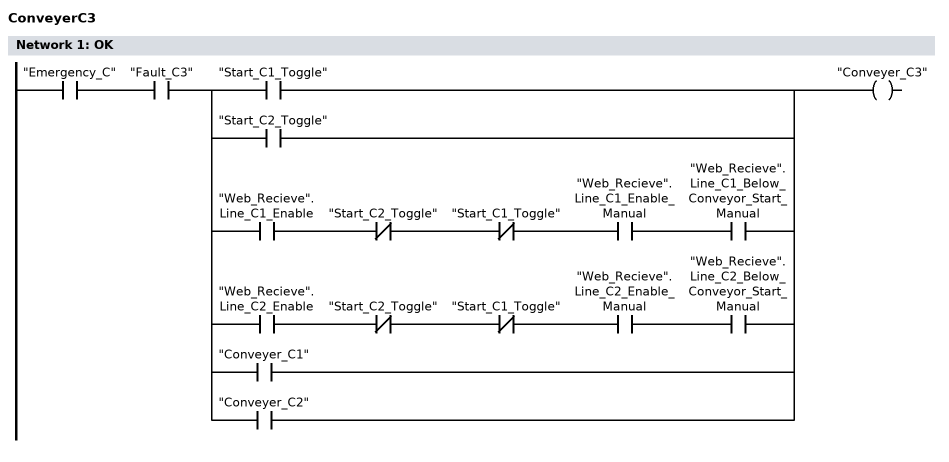
   RUNG wire#powerrail
      Contact( "Emergency_C" )
      Contact( "Fault_C3" )
      wire#w1
      Contact( "Start_C1_Toggle" )
      wire#w2
      Coil( "Conveyer_C3" )
   END_RUNG
   RUNG wire#w1
      Contact( "Start_C2_Toggle" )
   END_RUNG wire#w2
   RUNG wire#w1
      Contact( "Web_Recieve".Line_C1_Enable )
      I_Contact( "Start_C2_Toggle" )
      I_Contact( "Start_C1_Toggle" )
      Contact( "Web_Recieve".Line_C1_Enable_Manual )
      Contact( "Web_Recieve".Line_C1_Below_Conveyor_Start_Manual )
   END_RUNG wire#w2
   RUNG wire#w1
      Contact( "Web_Recieve".Line_C2_Enable )
      I_Contact( "Start_C2_Toggle" )
      I_Contact( "Start_C1_Toggle" )
      Contact( "Web_Recieve".Line_C2_Enable_Manual )
      Contact( "Web_Recieve".Line_C2_Below_Conveyor_Start_Manual )
   END_RUNG wire#w2
   RUNG wire#w1
      Contact( "Conveyer_C1" )
   END_RUNG wire#w2
   RUNG wire#w1
      Contact( "Conveyer_C2" )
   END_RUNG wire#w2
   // the same network as SCL:
   "Conveyer_C3" := "Emergency_C" AND "Fault_C3" AND ("Start_C1_Toggle" OR "Start_C2_Toggle" OR ("Web_Recieve".Line_C1_Enable AND NOT "Start_C2_Toggle" AND NOT "Start_C1_Toggle" AND "Web_Recieve".Line_C1_Enable_Manual AND "Web_Recieve".Line_C1_Below_Conveyor_Start_Manual) OR ("Web_Recieve".Line_C2_Enable AND NOT "Start_C2_Toggle" AND NOT "Start_C1_Toggle" AND "Web_Recieve".Line_C2_Enable_Manual AND "Web_Recieve".Line_C2_Below_Conveyor_Start_Manual) OR "Conveyer_C1" OR "Conveyer_C2");
END_REGION
END_FUNCTION_BLOCK

FUNCTION_BLOCK "WebDataPrepaare"   // FB10, SCL
{ S7_Optimized_Access := 'TRUE' }
VERSION : 0.1
BEGIN
   "Web_Send".C_Emergency := NOT "Emergency_C";
   "Web_Send".C1_Conveyer := "Conveyer_C1";
   "Web_Send".C2_Conveyer := "Conveyer_C2";
   "Web_Send".C3_Conveyor := "Conveyer_C3";

   "Web_Send".C1_Fault := NOT "Fault_C1";
   "Web_Send".C2_Fault := NOT "Fault_C2";
   "Web_Send".C3_Fault := NOT "Fault_C3";
   "Web_Send".C1_Silo_Low := "Low_Silo_C1";
   "Web_Send".C2_Silo_Low := "Low_Silo_C2";
   "Web_Send".C1_Silo_High := "HIgh_Silo_C1";
   "Web_Send".C2_Silo_High := "High_Silo_C2";
   "Web_Send".C1_Sample := "Pneumatic_C1";
   "Web_Send".C2_Sample := "Pneumatic_C2";
   "Web_Send".C1_Manual := "Web_Recieve".Line_C1_Enable_Manual;


   "Web_Send".C1_Running_Duration := "Web_Recieve".Line_C1_Conveyer_on_Time;
   "Web_Send".C1_Pause_Duration := "Web_Recieve".Line_C1_Conveyer_off_Time;
   "Web_Send".C1_Feeder_Vibration_Intensity := "Web_Recieve".Line_C1_Feeder_Intensity;
   "Web_Send".C1_Ruuning_Online := "Timer_On_C1_Conveyer".ET;
   "Web_Send".C1_Pause_Online := "Timer_Off_C1_Conveyer".ET;
   "Web_Send".C1_Sample_Interval :="Web_Recieve".Line_C1_Sampling_Time;
   "Web_Send".C1_Sample_Duration := "Web_Recieve".Line_C1_Sampling_OpenTime;
   "Web_Send".C1_Sample_Online := "Timer_Before_On_Sample_C1".ET - "Timer_Before_On_Sample_C1".ET;
   "Web_Send".C1_Enable := "Web_Recieve".Line_C1_Enable;
   "Web_Send".C1_Start := "Start_C1_Toggle";
   "Web_Send".C1_Empty_Line_Time := "Web_Recieve".Line_C1_Empty_Line_Time;
   "Web_Send".C1_Feeder_Delay_After_Start_Time := "Web_Recieve".Line_C1_Feeder_Delay_After_Start_Time;
   "Web_Send".C1_Feeder_Delay_Before_Stop_Time := "Web_Recieve".Line_C1_Feeder_Delay_Before_Stop_Time;
   "Web_Send".C1_Duration_Big_Silo_Stop_Time := "Web_Recieve".Line_C1_Big_Silo_Delay_Start;

   "Web_Send".C2_Running_Duration := "Web_Recieve".Line_C2_Conveyer_on_Time;
   "Web_Send".C2_Pause_Duration := "Web_Recieve".Line_C2_Conveyer_off_Time;
   "Web_Send".C2_Feeder_Vibration_Intensity := "Web_Recieve".Line_C2_Feeder_Intensity;
   "Web_Send".C2_Ruuning_Online := "Timer_On_C2_Conveyer".ET;
   "Web_Send".C2_Pause_Online := "Timer_Off_C2_Conveyer".ET;
   "Web_Send".C2_Sample_Interval := "Web_Recieve".Line_C2_Sampling_Time;
   "Web_Send".C2_Sample_Duration := "Web_Recieve".Line_C2_Sampling_OpenTime;
   "Web_Send".C2_Sample_Online := "Timer_Before_On_Sample_C2".ET - "Timer_Before_On_Sample_C2".ET;
   "Web_Send".C2_Enable := "Web_Recieve".Line_C2_Enable;
   "Web_Send".C2_Start := "Start_C2_Toggle";
   "Web_Send".C2_Empty_Line_Time := "Web_Recieve".Line_C2_Empty_Line_Time;
   "Web_Send".C2_Feeder_Delay_After_Start_Time := "Web_Recieve".Line_C2_Feeder_Delay_After_Start_Time;
   "Web_Send".C2_Feeder_Delay_Before_Stop_Time := "Web_Recieve".Line_C2_Feeder_Delay_Before_Stop_Time;
   "Web_Send".C2_Duration_Big_Silo_Stop_Time := "Web_Recieve".Line_C2_Big_Silo_Delay_Start;
END_FUNCTION_BLOCK

FUNCTION_BLOCK "Sample_C"   // FB11, LAD
{ S7_Optimized_Access := 'TRUE' }
VERSION : 0.1
   VAR_TEMP   // added for the SCL form of the ladder/FBD networks
      _w1 : Bool;
   END_VAR
BEGIN

REGION Network 1: C1 Before Sample
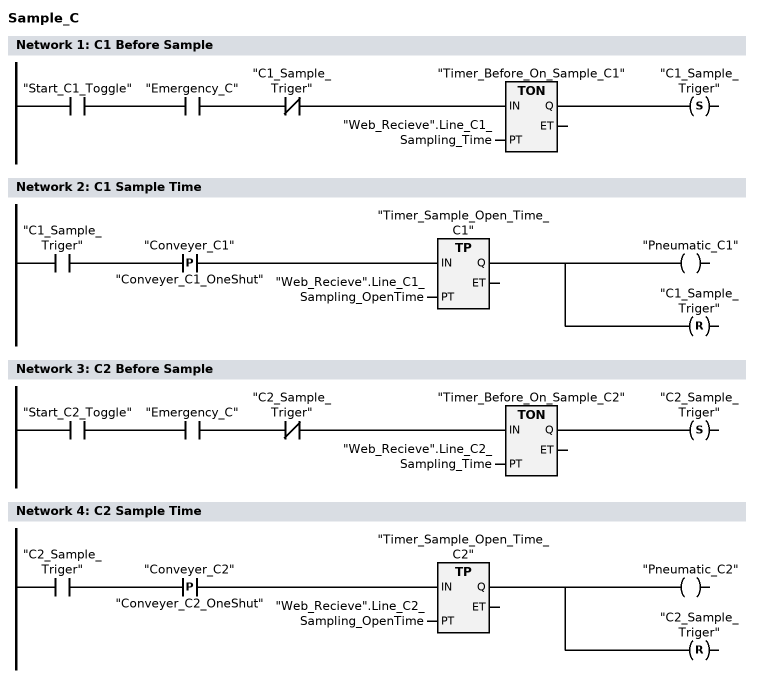
   "Timer_Before_On_Sample_C1".TON(IN := "Start_C1_Toggle" AND "Emergency_C" AND NOT "C1_Sample_Triger",
                           PT := "Web_Recieve".Line_C1_Sampling_Time);
   IF "Timer_Before_On_Sample_C1".Q THEN "C1_Sample_Triger" := TRUE; END_IF;
END_REGION

REGION Network 2: C1 Sample Time
   #_w1 := "C1_Sample_Triger" AND "Conveyer_C1" AND NOT "Conveyer_C1_OneShut";   // rising edge of "Conveyer_C1"
   "Conveyer_C1_OneShut" := "Conveyer_C1";
   "Timer_Sample_Open_Time_C1".TP(IN := #_w1, PT := "Web_Recieve".Line_C1_Sampling_OpenTime);
   "Pneumatic_C1" := "Timer_Sample_Open_Time_C1".Q;
   IF "Timer_Sample_Open_Time_C1".Q THEN "C1_Sample_Triger" := FALSE; END_IF;
END_REGION

REGION Network 3: C2 Before Sample
   "Timer_Before_On_Sample_C2".TON(IN := "Start_C2_Toggle" AND "Emergency_C" AND NOT "C2_Sample_Triger",
                           PT := "Web_Recieve".Line_C2_Sampling_Time);
   IF "Timer_Before_On_Sample_C2".Q THEN "C2_Sample_Triger" := TRUE; END_IF;
END_REGION

REGION Network 4: C2 Sample Time
   #_w1 := "C2_Sample_Triger" AND "Conveyer_C2" AND NOT "Conveyer_C2_OneShut";   // rising edge of "Conveyer_C2"
   "Conveyer_C2_OneShut" := "Conveyer_C2";
   "Timer_Sample_Open_Time_C2".TP(IN := #_w1, PT := "Web_Recieve".Line_C2_Sampling_OpenTime);
   "Pneumatic_C2" := "Timer_Sample_Open_Time_C2".Q;
   IF "Timer_Sample_Open_Time_C2".Q THEN "C2_Sample_Triger" := FALSE; END_IF;
END_REGION
END_FUNCTION_BLOCK

FUNCTION_BLOCK "Silo_Big_C"   // FB12, LAD
{ S7_Optimized_Access := 'TRUE' }
VERSION : 0.1
BEGIN

REGION Network 1
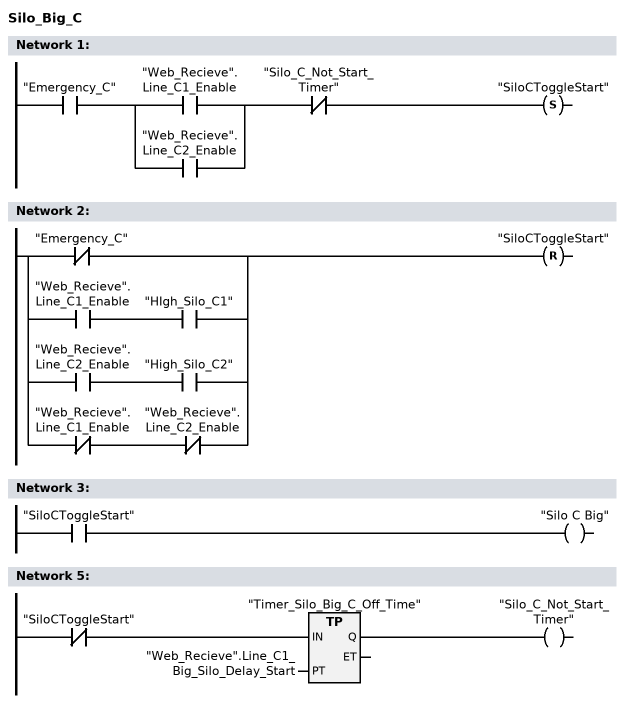
   RUNG wire#powerrail
      Contact( "Emergency_C" )
      wire#w1
      Contact( "Web_Recieve".Line_C1_Enable )
      wire#w2
      I_Contact( "Silo_C_Not_Start_Timer" )
      S_Coil( "SiloCToggleStart" )
   END_RUNG
   RUNG wire#w1
      Contact( "Web_Recieve".Line_C2_Enable )
   END_RUNG wire#w2
   // the same network as SCL:
   IF "Emergency_C" AND ("Web_Recieve".Line_C1_Enable OR "Web_Recieve".Line_C2_Enable) AND NOT "Silo_C_Not_Start_Timer" THEN
       "SiloCToggleStart" := TRUE;
   END_IF;
END_REGION

REGION Network 2
   RUNG wire#powerrail
      I_Contact( "Emergency_C" )
      wire#w1
      R_Coil( "SiloCToggleStart" )
   END_RUNG
   RUNG wire#powerrail
      Contact( "Web_Recieve".Line_C1_Enable )
      Contact( "HIgh_Silo_C1" )
   END_RUNG wire#w1
   RUNG wire#powerrail
      Contact( "Web_Recieve".Line_C2_Enable )
      Contact( "High_Silo_C2" )
   END_RUNG wire#w1
   RUNG wire#powerrail
      I_Contact( "Web_Recieve".Line_C1_Enable )
      I_Contact( "Web_Recieve".Line_C2_Enable )
   END_RUNG wire#w1
   // the same network as SCL:
   IF NOT "Emergency_C" OR ("Web_Recieve".Line_C1_Enable AND "HIgh_Silo_C1") OR ("Web_Recieve".Line_C2_Enable AND "High_Silo_C2") OR (NOT "Web_Recieve".Line_C1_Enable AND NOT "Web_Recieve".Line_C2_Enable) THEN
       "SiloCToggleStart" := FALSE;
   END_IF;
END_REGION

REGION Network 3
   RUNG wire#powerrail
      Contact( "SiloCToggleStart" )
      Coil( "Silo C Big" )
   END_RUNG
   // the same network as SCL:
   "Silo C Big" := "SiloCToggleStart";
END_REGION

REGION Network 5
   "Timer_Silo_Big_C_Off_Time".TP(IN := NOT "SiloCToggleStart",
                           PT := "Web_Recieve".Line_C1_Big_Silo_Delay_Start);
   "Silo_C_Not_Start_Timer" := "Timer_Silo_Big_C_Off_Time".Q;
END_REGION
END_FUNCTION_BLOCK

FUNCTION_BLOCK "Empty Line C1"   // FB13, LAD
{ S7_Optimized_Access := 'TRUE' }
VERSION : 0.1
BEGIN

REGION Network 1
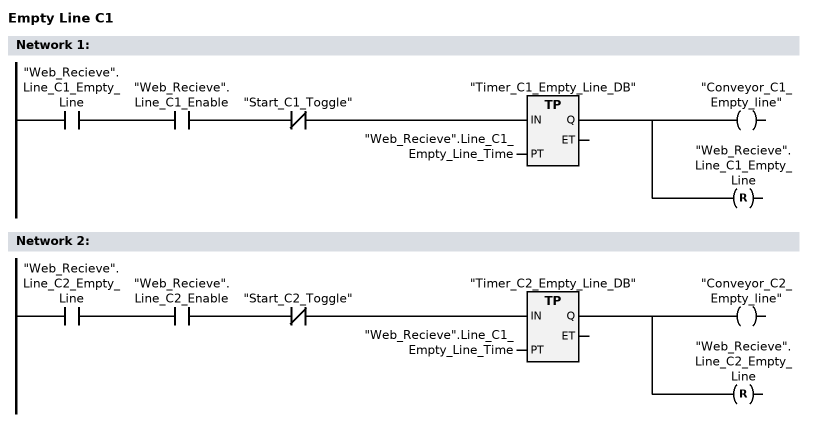
   "Timer_C1_Empty_Line_DB".TP(IN := "Web_Recieve".Line_C1_Empty_Line AND "Web_Recieve".Line_C1_Enable AND NOT "Start_C1_Toggle",
                           PT := "Web_Recieve".Line_C1_Empty_Line_Time);
   "Conveyor_C1_Empty_line" := "Timer_C1_Empty_Line_DB".Q;
   IF "Timer_C1_Empty_Line_DB".Q THEN "Web_Recieve".Line_C1_Empty_Line := FALSE; END_IF;
END_REGION

REGION Network 2
   "Timer_C2_Empty_Line_DB".TP(IN := "Web_Recieve".Line_C2_Empty_Line AND "Web_Recieve".Line_C2_Enable AND NOT "Start_C2_Toggle",
                           PT := "Web_Recieve".Line_C1_Empty_Line_Time);
   "Conveyor_C2_Empty_line" := "Timer_C2_Empty_Line_DB".Q;
   IF "Timer_C2_Empty_Line_DB".Q THEN "Web_Recieve".Line_C2_Empty_Line := FALSE; END_IF;
END_REGION
END_FUNCTION_BLOCK

ORGANIZATION_BLOCK "Main"   // OB1, LAD, ProgramCycle
TITLE = "Main Program Sweep (Cycle)"
{ S7_Optimized_Access := 'TRUE' }
VERSION : 0.1
   VAR_INPUT
      Initial_Call : Bool;   // Initial call of this OB
      Remanence : Bool;   // =True, if remanent data are available
   END_VAR
   VAR_TEMP
      TEMP : Int;
      clkRetVal : Int;
      newt : Int;
   END_VAR
BEGIN

REGION Network 1
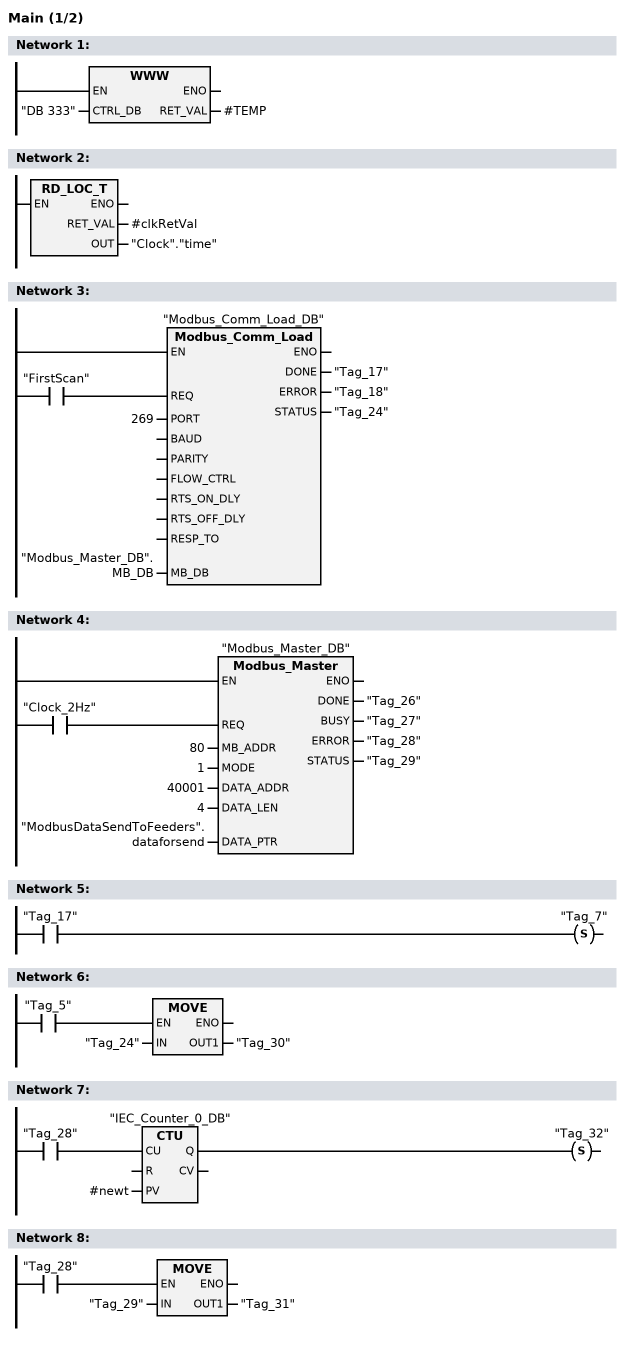
   #TEMP := WWW(CTRL_DB := "DB 333");
END_REGION

REGION Network 2
   #clkRetVal := RD_LOC_T(OUT => "Clock"."time");
END_REGION

REGION Network 3
   "Modbus_Comm_Load_DB"(REQ := "FirstScan",   // Modbus_Comm_Load
                         PORT := 269,
                         MB_DB := "Modbus_Master_DB".MB_DB,
                         DONE => "Tag_17",
                         ERROR => "Tag_18",
                         STATUS => "Tag_24");
END_REGION

REGION Network 4
   "Modbus_Master_DB"(REQ := "Clock_2Hz",   // Modbus_Master
                      MB_ADDR := 80,
                      MODE := 1,
                      DATA_ADDR := 40001,
                      DATA_LEN := 4,
                      DATA_PTR := "ModbusDataSendToFeeders".dataforsend,
                      DONE => "Tag_26",
                      BUSY => "Tag_27",
                      ERROR => "Tag_28",
                      STATUS => "Tag_29");
END_REGION

REGION Network 5
   RUNG wire#powerrail
      Contact( "Tag_17" )
      S_Coil( "Tag_7" )
   END_RUNG
   // the same network as SCL:
   IF "Tag_17" THEN "Tag_7" := TRUE; END_IF;
END_REGION

REGION Network 6
   RUNG wire#powerrail
      Contact( "Tag_5" )
      Move(in := "Tag_24", out1 => "Tag_30")
   END_RUNG
   // the same network as SCL:
   IF "Tag_5" THEN "Tag_30" := "Tag_24"; END_IF;
END_REGION

REGION Network 7
   "IEC_Counter_0_DB".CTU(CU := "Tag_28", PV := #newt);
   IF "IEC_Counter_0_DB".Q THEN "Tag_32" := TRUE; END_IF;
END_REGION

REGION Network 8
   RUNG wire#powerrail
      Contact( "Tag_28" )
      Move(in := "Tag_29", out1 => "Tag_31")
   END_RUNG
   // the same network as SCL:
   IF "Tag_28" THEN "Tag_31" := "Tag_29"; END_IF;
END_REGION

REGION Network 9
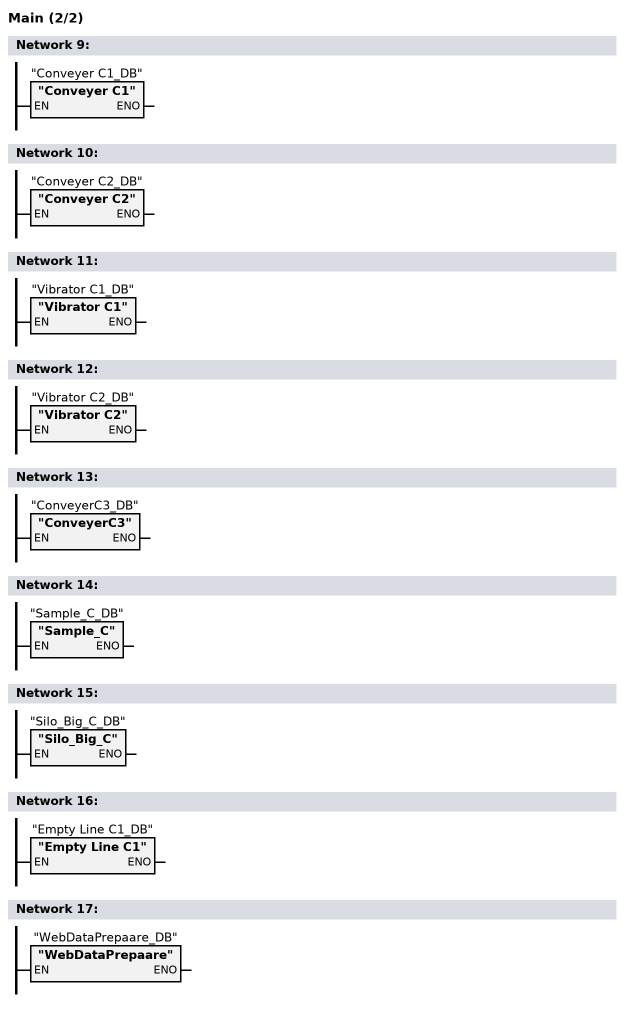
   RUNG wire#powerrail
      "Conveyer C1_DB"()
   END_RUNG
   // the same network as SCL:
   "Conveyer C1_DB"();   // "Conveyer C1"
END_REGION

REGION Network 10
   RUNG wire#powerrail
      "Conveyer C2_DB"()
   END_RUNG
   // the same network as SCL:
   "Conveyer C2_DB"();   // "Conveyer C2"
END_REGION

REGION Network 11
   RUNG wire#powerrail
      "Vibrator C1_DB"()
   END_RUNG
   // the same network as SCL:
   "Vibrator C1_DB"();   // "Vibrator C1"
END_REGION

REGION Network 12
   RUNG wire#powerrail
      "Vibrator C2_DB"()
   END_RUNG
   // the same network as SCL:
   "Vibrator C2_DB"();   // "Vibrator C2"
END_REGION

REGION Network 13
   RUNG wire#powerrail
      "ConveyerC3_DB"()
   END_RUNG
   // the same network as SCL:
   "ConveyerC3_DB"();   // "ConveyerC3"
END_REGION

REGION Network 14
   RUNG wire#powerrail
      "Sample_C_DB"()
   END_RUNG
   // the same network as SCL:
   "Sample_C_DB"();   // "Sample_C"
END_REGION

REGION Network 15
   RUNG wire#powerrail
      "Silo_Big_C_DB"()
   END_RUNG
   // the same network as SCL:
   "Silo_Big_C_DB"();   // "Silo_Big_C"
END_REGION

REGION Network 16
   RUNG wire#powerrail
      "Empty Line C1_DB"()
   END_RUNG
   // the same network as SCL:
   "Empty Line C1_DB"();   // "Empty Line C1"
END_REGION

REGION Network 17
   RUNG wire#powerrail
      "WebDataPrepaare_DB"()
   END_RUNG
   // the same network as SCL:
   "WebDataPrepaare_DB"();   // "WebDataPrepaare"
END_REGION
END_ORGANIZATION_BLOCK

// ===== PLC "PLC_1"  CPU 1516-3 PN/DP =====

VAR_GLOBAL   // PLC tag table "Default tag table"
   "Tag_31" AT %M100.5 : Bool;
   "Run consent OS" AT %M151.6 : Bool;
   "Run_Consent_A1_Negetive_OS" AT %M151.7 : Bool;
   "Vibrator_A2_Remaning_Time" AT %MD166 : DInt;
   "System_Byte(1)" AT %MB1 : Byte;
   "FirstScan" AT %M1.0 : Bool;
END_VAR

VAR_GLOBAL   // PLC tag table "Default tag table_1"
   "Phase_Control" AT %I8.0 : Bool;
   "Start_A" AT %I8.7 : Bool;
   "Spare_6" AT %I9.6 : Bool;
   "Spare_7" AT %I9.7 : Bool;
   "Emergency_A" AT %I8.4 : Bool;
   "Fault_A1" AT %I8.1 : Bool;
   "Low_Silo_A1" AT %I0.2 : Bool;
   "Low_Silo_A2" AT %I0.1 : Bool;
   "Low_Silo_B1" AT %I0.7 : Bool;
   "Low_Silo_B2" AT %I0.4 : Bool;
   "High_Silo_A1" AT %I0.3 : Bool;
   "High_Silo_A2" AT %I0.0 : Bool;
   "High_Silo_B1" AT %I0.6 : Bool;
   "High_Silo_B2" AT %I0.5 : Bool;
   "Fault_A2" AT %I9.1 : Bool;
   "Fault_B1" AT %I8.2 : Bool;
   "Fault_B2" AT %I9.2 : Bool;
   "Fault_A3" AT %I9.5 : Bool;
   "Fault_B3" AT %I9.4 : Bool;
   "Emergency_B" AT %I9.3 : Bool;
   "Rel Spare_4" AT %Q2.4 : Bool;
   "Rel Spare_5" AT %Q2.5 : Bool;
   "Rel Spare_6" AT %Q2.6 : Bool;
   "Rel Spare_7" AT %Q2.7 : Bool;
   "Rel Spare_8" AT %Q3.0 : Bool;
   "Rel Spare_9" AT %Q3.1 : Bool;
   "Rel Spare_10" AT %Q3.2 : Bool;
   "Rel Spare_11" AT %Q3.3 : Bool;
   "Rel Spare_12" AT %Q3.4 : Bool;
   "Rel Spare_13" AT %Q3.5 : Bool;
   "Rel Spare_14" AT %Q3.6 : Bool;
   "Rel Spare_15" AT %Q3.7 : Bool;
   "Light_A1" AT %Q2.3 : Bool;
   "Light_A2" AT %Q2.2 : Bool;
   "Light_B1" AT %Q2.1 : Bool;
   "Light_B2" AT %Q2.0 : Bool;
   "Conveyer_A1" AT %Q0.4 : Bool;
   "Conveyer_A2" AT %Q0.5 : Bool;
   "Conveyer_B1" AT %Q9.0 : Bool;
   "Conveyer_B2" AT %Q8.0 : Bool;
   "Pneumatic_A1" AT %Q9.1 : Bool;
   "Pneumatic_A2" AT %Q8.1 : Bool;
   "Pneumatic_B1" AT %Q8.2 : Bool;
   "Pneumatic_B2" AT %Q9.2 : Bool;
   "Conveyer_A3" AT %Q9.5 : Bool;
   "Conveyer_B3_Left" AT %Q9.6 : Bool;
   "Conveyer_B3_Right" AT %Q8.5 : Bool;
   "Tag_1(1)" AT %M10.0 : Bool;
   "Tag_2" AT %M10.1 : Bool;
   "start" AT %M10.2 : Bool;
   "Tag_3" AT %M110.0 : Bool;
   "Tag_10" AT %M110.1 : Bool;
   "Tag_11" AT %M110.2 : Bool;
   "System_Byte" AT %MB1 : Byte;
   "DiagStatusUpdate" AT %M1.1 : Bool;
   "AlwaysTRUE" AT %M1.2 : Bool;
   "AlwaysFALSE" AT %M1.3 : Bool;
   "Clock_Byte" AT %MB0 : Byte;
   "Clock_10Hz" AT %M0.0 : Bool;
   "Clock_5Hz" AT %M0.1 : Bool;
   "Clock_2.5Hz" AT %M0.2 : Bool;
   "Clock_2Hz" AT %M0.3 : Bool;
   "Clock_1.25Hz" AT %M0.4 : Bool;
   "Clock_1Hz" AT %M0.5 : Bool;
   "Clock_0.625Hz" AT %M0.6 : Bool;
   "Clock_0.5Hz" AT %M0.7 : Bool;
   "Tag_12" AT %M120.1 : Bool;
   "Tag_13" AT %M120.0 : Bool;
   "Tag_14" AT %M120.2 : Bool;
   "Tag_15" AT %MW112 : Word;
   "Tag_16" AT %MW114 : Word;
   "Tag_17" AT %MW122 : Word;
   "Tag_18" AT %MW124 : Word;
   "Tag_4" AT %M1000.0 : Bool;
   "Tag_5" AT %M1000.1 : Bool;
   "Tag_6" AT %MW1002 : Word;
   "Tag_7" AT %M1000.4 : Bool;
   "Tag_8" AT %MW1004 : Word;
   "Tag_9" AT %M1010.0 : Bool;
   "Tag_19" AT %M1010.1 : Bool;
   "Tag_20" AT %M1010.2 : Bool;
   "Tag_21" AT %MW1012 : Word;
   "Tag_22" AT %M1010.4 : Bool;
   "Tag_23" AT %MW1014 : Word;
   "Tag_24" AT %M990.0 : Bool;
   "Tag_25" AT %M990.5 : Bool;
   "Line_A1_Start_Consent" AT %M150.0 : Bool;
   "Line_A1_Run_Consent" AT %M150.1 : Bool;
   "Line_A1_Conveyer_Timer" AT %M150.2 : Bool;
   "A1_Start_Conveyer" AT %M150.3 : Bool;
   "TriggerStartToggleMemory" AT %M150.4 : Bool;
   "Start_A1_Toggle" AT %M150.5 : Bool;
   "TriggerA1ToggleStop" AT %M150.6 : Bool;
   "Conveyer_A1_On" AT %M150.7 : Bool;
   "Conveyer_A1_Off" AT %M151.0 : Bool;
   "Line_A2_Start_Consent" AT %M160.0 : Bool;
   "Line_A2_Run_Consent" AT %M160.1 : Bool;
   "Line_A2_Conveyer_Timer" AT %M160.2 : Bool;
   "A2_Start_Conveyer" AT %M160.3 : Bool;
   "TriggerStopToggleMemoryA2" AT %M160.6 : Bool;
   "TriggerStartToggleMemoryA2" AT %M160.4 : Bool;
   "Start_A2_Toggle" AT %M160.5 : Bool;
   "Conveyer_A2_Off" AT %M161.0 : Bool;
   "Conveyer_A2_On" AT %M160.7 : Bool;
   "Line_B1_Start_Consent" AT %M170.0 : Bool;
   "Line_B1_Run_Consent" AT %M170.1 : Bool;
   "Line_B1_Conveyer_Timer" AT %M170.2 : Bool;
   "B1_Start_Conveyer" AT %M170.3 : Bool;
   "Start_B1_Toggle" AT %M170.5 : Bool;
   "TriggerStartToggleMemoryB1" AT %M170.4 : Bool;
   "TriggerB1ToggleStop" AT %M170.6 : Bool;
   "Conveyer_B1_Off" AT %M171.0 : Bool;
   "Conveyer_B1_On" AT %M170.7 : Bool;
   "Line_B2_Start_Consent" AT %M180.0 : Bool;
   "Line_B2_Run_Consent" AT %M180.1 : Bool;
   "B2_Start_Conveyer" AT %M180.3 : Bool;
   "Line_B2_Conveyer_Timer" AT %M180.2 : Bool;
   "Start_B2_Toggle" AT %M180.5 : Bool;
   "TriggerStartToggleMemoryB2" AT %M180.4 : Bool;
   "TriggerStopToggleMemoryB2" AT %M180.6 : Bool;
   "Conveyer_B2_Off" AT %M181.0 : Bool;
   "Conveyer_B2_On" AT %M180.7 : Bool;
   "Vibrator_A1_On" AT %M151.4 : Bool;
   "Vibrator_A2_On" AT %M161.4 : Bool;
   "Vibrator_B1_On" AT %M171.4 : Bool;
   "Vibrator_B2_On" AT %M181.4 : Bool;
   "A1_Sample_Triger" AT %M151.1 : Bool;
   "Conveyer_A1_OneShut" AT %M151.2 : Bool;
   "Tag_27" AT %M151.3 : Bool;
   "A2_Sample_Triger" AT %M161.1 : Bool;
   "Conveyer_A2_OneShut" AT %M161.2 : Bool;
   "B1_Sample_Triger" AT %M171.1 : Bool;
   "Conveyer_B1_OneShut" AT %M171.2 : Bool;
   "B2_Sample_Triger" AT %M181.1 : Bool;
   "Conveyer_B2_OneShut" AT %M181.2 : Bool;
   "B_Emergency_Flag" AT %M171.3 : Bool;
   "SiloAToggleStart" AT %M190.0 : Bool;
   "SiloBToggleStart" AT %M190.1 : Bool;
   "Conveyor_B3_Left" AT %M200.0 : Bool;
   "Conveyor_B3_Right" AT %M200.1 : Bool;
   "Silo_B_Not_Start_Timer" AT %M190.3 : Bool;
   "Silo_A_Not_Start_Timer" AT %M190.2 : Bool;
   "Conveyor_B3_Start" AT %M190.4 : Bool;
   "Conveyor_A1_Empty_line" AT %M151.5 : Bool;
   "Conveyor_A2_Empty_line" AT %M161.5 : Bool;
   "Conveyor_B1_Empty_line" AT %M171.5 : Bool;
   "Conveyor_B2_Empty_line" AT %M181.5 : Bool;
   "Vibrator_A1_Remaning_Time" AT %MD156 : DInt;
   "Tag_29" AT %MD176 : DInt;
   "Tag_30" AT %MD186 : DInt;
END_VAR

VAR_GLOBAL CONSTANT   // PLC tag table "Default tag table_1"
   "None(1)" : Pip := 65535;
   "Automatic update(1)" : Pip := 0;
   "PIP 1(1)" : Pip := 1;
   "PIP 2(1)" : Pip := 2;
   "PIP 3(1)" : Pip := 3;
   "PIP 4(1)" : Pip := 4;
   "PIP OB Servo(1)" : Pip := 32768;
   "Local~MC(1)" : Hw_SubModule := 51;
   "Local~Common(1)" : Hw_SubModule := 50;
   "Local~Device(1)" : Hw_Device := 32;
   "Local~Configuration(1)" : Hw_SubModule := 33;
   "Local~Exec(1)" : Hw_SubModule := 52;
   "Local(1)" : Hw_SubModule := 49;
   "Local~PROFINET_interface_1(1)" : Hw_Interface := 64;
   "Local~PROFINET_interface_1~Port_1(1)" : Hw_Interface := 65;
   "Local~HSC_1" : Hw_Hsc := 257;
   "Local~HSC_2" : Hw_Hsc := 258;
   "Local~HSC_3" : Hw_Hsc := 259;
   "Local~HSC_4" : Hw_Hsc := 260;
   "Local~HSC_5" : Hw_Hsc := 261;
   "Local~HSC_6" : Hw_Hsc := 262;
   "Local~AI_2_1" : Hw_SubModule := 263;
   "Local~DI_8_DQ_6_1" : Hw_SubModule := 264;
   "Local~Pulse_1" : Hw_Pwm := 265;
   "Local~Pulse_2" : Hw_Pwm := 266;
   "Local~Pulse_3" : Hw_Pwm := 267;
   "Local~Pulse_4" : Hw_Pwm := 268;
   "Local~CB_1241_(RS485)" : Port := 269;
   "Local~DQ_16xRelay_1" : Hw_SubModule := 270;
   "Local~DI_16x24VDC_DQ_16xRelay_1" : Hw_SubModule := 271;
   "OB_Main(1)" : OB_PCYCLE := 1;
END_VAR

DATA_BLOCK "ScenarioData"   // DB1
{ S7_Optimized_Access := 'TRUE' }
VERSION : 0.1
   VAR
      DefaultScenario : Int := 1;
      Line_A1_Conveyer_on_Time_Scenario_A : DInt := 2;
      Line_A1_Conveyer_off_Time_Scenario_A : DInt := 3;
      Line_A1_Sampling_Time_Scenario_A : DInt := 4;
      Line_A1_Sampling_OpenTime_Scenario_A : DInt := 5;
      Line_A1_Feeder_Intensity_Scenario_A : Int := 6;
      Line_A1_Duration_Big_Silo_Off_Scenario_A : DInt := 7;
      Line_A1_Feeder_Delay_Before_Stop_Time_Scenario_A : DInt := 8;
      Line_A1_Feeder_Delay_After_Start_Time_Scenario_A : DInt := 9;
      Line_A1_Conveyer_on_Time_Scenario_B : DInt := 10;
      Line_A1_Conveyer_off_Time_Scenario_B : DInt := 11;
      Line_A1_Sampling_Time_Scenario_B : DInt := 12;
      Line_A1_Sampling_OpenTime_Scenario_B : DInt := 13;
      Line_A1_Feeder_Intensity_Scenario_B : Int := 14;
      Line_A1_Duration_Big_Silo_Off_Scenario_B : DInt := 15;
      Line_A1_Feeder_Delay_Before_Stop_Time_Scenario_B : DInt := 16;
      Line_A1_Feeder_Delay_After_Start_Time_Scenario_B : DInt := 17;
      Line_A1_Conveyer_on_Time_Scenario_C : DInt := 18;
      Line_A1_Conveyer_off_Time_Scenario_C : DInt := 19;
      Line_A1_Sampling_Time_Scenario_C : DInt := 20;
      Line_A1_Sampling_OpenTime_Scenario_C : DInt := 21;
      Line_A1_Feeder_Intensity_Scenario_C : Int := 22;
      Line_A1_Duration_Big_Silo_Off_Scenario_C : DInt := 23;
      Line_A1_Feeder_Delay_Before_Stop_Time_Scenario_C : DInt := 24;
      Line_A1_Feeder_Delay_After_Start_Time_Scenario_C : DInt := 25;
      Line_A1_Conveyer_on_Time_Scenario_E : DInt := 26;
      Line_A1_Conveyer_off_Time_Scenario_E : DInt := 27;
      Line_A1_Sampling_Time_Scenario_E : DInt := 28;
      Line_A1_Sampling_OpenTime_Scenario_E : DInt := 29;
      Line_A1_Feeder_Intensity_Scenario_E : Int := 30;
      Line_A1_Duration_Big_Silo_Off_Scenario_E : DInt := 31;
      Line_A1_Feeder_Delay_Before_Stop_Time_Scenario_E : DInt := 32;
      Line_A1_Feeder_Delay_After_Start_Time_Scenario_E : DInt := 33;
      Line_A1_Conveyer_on_Time_Scenario_D : DInt := 34;
      Line_A1_Conveyer_off_Time_Scenario_D : DInt := 35;
      Line_A1_Sampling_Time_Scenario_D : DInt := 36;
      Line_A1_Sampling_OpenTime_Scenario_D : DInt := 37;
      Line_A1_Feeder_Intensity_Scenario_D : Int := 38;
      Line_A1_Duration_Big_Silo_Off_Scenario_D : DInt := 39;
      Line_A1_Feeder_Delay_Before_Stop_Time_Scenario_D : DInt := 40;
      Line_A1_Feeder_Delay_After_Start_Time_Scenario_D : DInt := 41;
      Line_A2_Conveyer_on_Time_Scenario_A : DInt := 42;
      Line_A2_Conveyer_off_Time_Scenario_A : DInt := 43;
      Line_A2_Sampling_Time_Scenario_A : DInt := 44;
      Line_A2_Sampling_OpenTime_Scenario_A : DInt := 45;
      Line_A2_Feeder_Intensity_Scenario_A : Int := 46;
      Line_A2_Duration_Big_Silo_Off_Scenario_A : DInt := 47;
      Line_A2_Feeder_Delay_Before_Stop_Time_Scenario_A : DInt := 48;
      Line_A2_Feeder_Delay_After_Start_Time_Scenario_A : DInt := 49;
      Line_A2_Conveyer_on_Time_Scenario_B : DInt := 50;
      Line_A2_Conveyer_off_Time_Scenario_B : DInt := 51;
      Line_A2_Sampling_Time_Scenario_B : DInt := 52;
      Line_A2_Sampling_OpenTime_Scenario_B : DInt := 53;
      Line_A2_Feeder_Intensity_Scenario_B : Int := 54;
      Line_A2_Duration_Big_Silo_Off_Scenario_B : DInt := 55;
      Line_A2_Feeder_Delay_Before_Stop_Time_Scenario_B : DInt := 56;
      Line_A2_Feeder_Delay_After_Start_Time_Scenario_B : DInt := 57;
      Line_A2_Conveyer_on_Time_Scenario_C : DInt := 58;
      Line_A2_Conveyer_off_Time_Scenario_C : DInt := 59;
      Line_A2_Sampling_Time_Scenario_C : DInt := 60;
      Line_A2_Sampling_OpenTime_Scenario_C : DInt := 61;
      Line_A2_Feeder_Intensity_Scenario_C : Int := 62;
      Line_A2_Duration_Big_Silo_Off_Scenario_C : DInt := 63;
      Line_A2_Feeder_Delay_Before_Stop_Time_Scenario_C : DInt := 64;
      Line_A2_Feeder_Delay_After_Start_Time_Scenario_C : DInt := 65;
      Line_A2_Conveyer_on_Time_Scenario_E : DInt := 66;
      Line_A2_Conveyer_off_Time_Scenario_E : DInt := 67;
      Line_A2_Sampling_Time_Scenario_E : DInt := 68;
      Line_A2_Sampling_OpenTime_Scenario_E : DInt := 69;
      Line_A2_Feeder_Intensity_Scenario_E : Int := 70;
      Line_A2_Duration_Big_Silo_Off_Scenario_E : DInt := 71;
      Line_A2_Feeder_Delay_Before_Stop_Time_Scenario_E : DInt := 72;
      Line_A2_Feeder_Delay_After_Start_Time_Scenario_E : DInt := 73;
      Line_A2_Conveyer_on_Time_Scenario_D : DInt := 74;
      Line_A2_Conveyer_off_Time_Scenario_D : DInt := 75;
      Line_A2_Sampling_Time_Scenario_D : DInt := 76;
      Line_A2_Sampling_OpenTime_Scenario_D : DInt := 77;
      Line_A2_Feeder_Intensity_Scenario_D : Int := 78;
      Line_A2_Duration_Big_Silo_Off_Scenario_D : DInt := 79;
      Line_A2_Feeder_Delay_Before_Stop_Time_Scenario_D : DInt := 80;
      Line_A2_Feeder_Delay_After_Start_Time_Scenario_D : DInt := 81;
      Line_B1_Conveyer_on_Time_Scenario_A : DInt := 82;
      Line_B1_Conveyer_off_Time_Scenario_A : DInt := 83;
      Line_B1_Sampling_Time_Scenario_A : DInt := 84;
      Line_B1_Sampling_OpenTime_Scenario_A : DInt := 85;
      Line_B1_Feeder_Intensity_Scenario_A : Int := 86;
      Line_B1_Duration_Big_Silo_Off_Scenario_A : DInt := 87;
      Line_B1_Feeder_Delay_Before_Stop_Time_Scenario_A : DInt := 88;
      Line_B1_Feeder_Delay_After_Start_Time_Scenario_A : DInt := 89;
      Line_B1_Conveyer_on_Time_Scenario_B : DInt := 90;
      Line_B1_Conveyer_off_Time_Scenario_B : DInt := 91;
      Line_B1_Sampling_Time_Scenario_B : DInt := 92;
      Line_B1_Sampling_OpenTime_Scenario_B : DInt := 93;
      Line_B1_Feeder_Intensity_Scenario_B : Int := 94;
      Line_B1_Duration_Big_Silo_Off_Scenario_B : DInt := 95;
      Line_B1_Feeder_Delay_Before_Stop_Time_Scenario_B : DInt := 96;
      Line_B1_Feeder_Delay_After_Start_Time_Scenario_B : DInt := 97;
      Line_B1_Conveyer_on_Time_Scenario_C : DInt := 98;
      Line_B1_Conveyer_off_Time_Scenario_C : DInt := 99;
      Line_B1_Sampling_Time_Scenario_C : DInt := 100;
      Line_B1_Sampling_OpenTime_Scenario_C : DInt := 101;
      Line_B1_Feeder_Intensity_Scenario_C : Int := 102;
      Line_B1_Duration_Big_Silo_Off_Scenario_C : DInt := 103;
      Line_B1_Feeder_Delay_Before_Stop_Time_Scenario_C : DInt := 104;
      Line_B1_Feeder_Delay_After_Start_Time_Scenario_C : DInt := 105;
      Line_B1_Conveyer_on_Time_Scenario_E : DInt := 106;
      Line_B1_Conveyer_off_Time_Scenario_E : DInt := 107;
      Line_B1_Sampling_Time_Scenario_E : DInt := 108;
      Line_B1_Sampling_OpenTime_Scenario_E : DInt := 109;
      Line_B1_Feeder_Intensity_Scenario_E : Int := 110;
      Line_B1_Duration_Big_Silo_Off_Scenario_E : DInt := 111;
      Line_B1_Feeder_Delay_Before_Stop_Time_Scenario_E : DInt := 112;
      Line_B1_Feeder_Delay_After_Start_Time_Scenario_E : DInt := 113;
      Line_B1_Conveyer_on_Time_Scenario_D : DInt := 114;
      Line_B1_Conveyer_off_Time_Scenario_D : DInt := 115;
      Line_B1_Sampling_Time_Scenario_D : DInt := 116;
      Line_B1_Sampling_OpenTime_Scenario_D : DInt := 117;
      Line_B1_Feeder_Intensity_Scenario_D : Int := 118;
      Line_B1_Duration_Big_Silo_Off_Scenario_D : DInt := 119;
      Line_B1_Feeder_Delay_Before_Stop_Time_Scenario_D : DInt := 120;
      Line_B1_Feeder_Delay_After_Start_Time_Scenario_D : DInt := 121;
      Line_B2_Conveyer_on_Time_Scenario_A : DInt := 122;
      Line_B2_Conveyer_off_Time_Scenario_A : DInt := 123;
      Line_B2_Sampling_Time_Scenario_A : DInt := 124;
      Line_B2_Sampling_OpenTime_Scenario_A : DInt := 125;
      Line_B2_Feeder_Intensity_Scenario_A : Int := 126;
      Line_B2_Duration_Big_Silo_Off_Scenario_A : DInt := 127;
      Line_B2_Feeder_Delay_Before_Stop_Time_Scenario_A : DInt := 128;
      Line_B2_Feeder_Delay_After_Start_Time_Scenario_A : DInt := 129;
      Line_B2_Conveyer_on_Time_Scenario_B : DInt := 130;
      Line_B2_Conveyer_off_Time_Scenario_B : DInt := 131;
      Line_B2_Sampling_Time_Scenario_B : DInt := 132;
      Line_B2_Sampling_OpenTime_Scenario_B : DInt := 133;
      Line_B2_Feeder_Intensity_Scenario_B : Int := 134;
      Line_B2_Duration_Big_Silo_Off_Scenario_B : DInt := 135;
      Line_B2_Feeder_Delay_Before_Stop_Time_Scenario_B : DInt := 136;
      Line_B2_Feeder_Delay_After_Start_Time_Scenario_B : DInt := 137;
      Line_B2_Conveyer_on_Time_Scenario_C : DInt := 138;
      Line_B2_Conveyer_off_Time_Scenario_C : DInt := 139;
      Line_B2_Sampling_Time_Scenario_C : DInt := 140;
      Line_B2_Sampling_OpenTime_Scenario_C : DInt := 141;
      Line_B2_Feeder_Intensity_Scenario_C : Int := 142;
      Line_B2_Duration_Big_Silo_Off_Scenario_C : DInt := 143;
      Line_B2_Feeder_Delay_Before_Stop_Time_Scenario_C : DInt := 144;
      Line_B2_Feeder_Delay_After_Start_Time_Scenario_C : DInt := 145;
      Line_B2_Conveyer_on_Time_Scenario_E : DInt := 146;
      Line_B2_Conveyer_off_Time_Scenario_E : DInt := 147;
      Line_B2_Sampling_Time_Scenario_E : DInt := 148;
      Line_B2_Sampling_OpenTime_Scenario_E : DInt := 149;
      Line_B2_Feeder_Intensity_Scenario_E : Int := 150;
      Line_B2_Duration_Big_Silo_Off_Scenario_E : DInt := 151;
      Line_B2_Feeder_Delay_Before_Stop_Time_Scenario_E : DInt := 152;
      Line_B2_Feeder_Delay_After_Start_Time_Scenario_E : DInt := 153;
      Line_B2_Conveyer_on_Time_Scenario_D : DInt := 154;
      Line_B2_Conveyer_off_Time_Scenario_D : DInt := 155;
      Line_B2_Sampling_Time_Scenario_D : DInt := 156;
      Line_B2_Sampling_OpenTime_Scenario_D : DInt := 157;
      Line_B2_Feeder_Intensity_Scenario_D : Int := 158;
      Line_B2_Duration_Big_Silo_Off_Scenario_D : DInt := 159;
      Line_B2_Feeder_Delay_Before_Stop_Time_Scenario_D : DInt := 160;
      Line_B2_Feeder_Delay_After_Start_Time_Scenario_D : DInt := 161;
      Line_A1_Empty_Line_Time_Scenario_A : DInt := 162;
      Line_A2_Empty_Line_Time_Scenario_A : DInt := 163;
      Line_B1_Empty_Line_Time_Scenario_A : DInt := 164;
      Line_B2_Empty_Line_Time_Scenario_A : DInt := 165;
      Line_A1_Empty_Line_Time_Scenario_B : DInt := 166;
      Line_A2_Empty_Line_Time_Scenario_B : DInt := 167;
      Line_B1_Empty_Line_Time_Scenario_B : DInt := 168;
      Line_B2_Empty_Line_Time_Scenario_B : DInt := 169;
      Line_A1_Empty_Line_Time_Scenario_C : DInt := 170;
      Line_A2_Empty_Line_Time_Scenario_C : DInt := 171;
      Line_B1_Empty_Line_Time_Scenario_C : DInt := 172;
      Line_B2_Empty_Line_Time_Scenario_C : DInt := 173;
      Line_A1_Empty_Line_Time_Scenario_D : DInt := 174;
      Line_A2_Empty_Line_Time_Scenario_D : DInt := 175;
      Line_B1_Empty_Line_Time_Scenario_D : DInt := 176;
      Line_B2_Empty_Line_Time_Scenario_D : DInt := 177;
      Line_A1_Empty_Line_Time_Scenario_E : DInt := 178;
      Line_A2_Empty_Line_Time_Scenario_E : DInt := 179;
      Line_B1_Empty_Line_Time_Scenario_E : DInt := 180;
      Line_B2_Empty_Line_Time_Scenario_E : DInt := 181;
   END_VAR
BEGIN
END_DATA_BLOCK

DATA_BLOCK "Conveyer B1_DB"   // DB3
{ S7_Optimized_Access := 'TRUE' }
VERSION : 0.1
// stored: InstanceOfName Conveyer B1
"Conveyer B1"
BEGIN
END_DATA_BLOCK

DATA_BLOCK "ModbusDataSendToFeeders"   // DB7
{ S7_Optimized_Access := 'FALSE' }
VERSION : 0.1
   VAR
      dataforsend : Array[0..3] of Int;
   END_VAR
BEGIN
   dataforsend[0] := 0;
   dataforsend[1] := 0;
   dataforsend[2] := 0;
   dataforsend[3] := 0;
END_DATA_BLOCK

DATA_BLOCK "Conveyer A1_DB"   // DB12
{ S7_Optimized_Access := 'TRUE' }
VERSION : 0.1
// stored: InstanceOfName Conveyer A1
"Conveyer A1"
BEGIN
END_DATA_BLOCK

DATA_BLOCK "Conveyer A2_DB"   // DB13
{ S7_Optimized_Access := 'TRUE' }
VERSION : 0.1
// stored: InstanceOfName Conveyer A2
"Conveyer A2"
BEGIN
END_DATA_BLOCK

DATA_BLOCK "Conveyer B1_DB_1"   // DB17
{ S7_Optimized_Access := 'TRUE' }
VERSION : 0.1
// stored: InstanceOfName Conveyer B1
"Conveyer B1"
BEGIN
END_DATA_BLOCK

DATA_BLOCK "Conveyer B2_DB"   // DB18
{ S7_Optimized_Access := 'TRUE' }
VERSION : 0.1
// stored: InstanceOfName Conveyer B2
"Conveyer B2"
BEGIN
END_DATA_BLOCK

DATA_BLOCK "Vibrator A1_DB"   // DB19
{ S7_Optimized_Access := 'TRUE' }
VERSION : 0.1
// stored: InstanceOfName Vibrator A1
"Vibrator A1"
BEGIN
END_DATA_BLOCK

DATA_BLOCK "Vibrator A2_DB"   // DB20
{ S7_Optimized_Access := 'TRUE' }
VERSION : 0.1
// stored: InstanceOfName Vibrator A2
"Vibrator A2"
BEGIN
END_DATA_BLOCK

DATA_BLOCK "Vibrator B1_DB"   // DB21
{ S7_Optimized_Access := 'TRUE' }
VERSION : 0.1
// stored: InstanceOfName Vibrator B1
"Vibrator B1"
BEGIN
END_DATA_BLOCK

DATA_BLOCK "Vibrator B2_DB"   // DB22
{ S7_Optimized_Access := 'TRUE' }
VERSION : 0.1
// stored: InstanceOfName Vibrator B2
"Vibrator B2"
BEGIN
END_DATA_BLOCK

DATA_BLOCK "Web_Send"   // DB23
{ S7_Optimized_Access := 'TRUE' }
VERSION : 0.1
   VAR
      "time" : DTL;
      ModbusDone : Bool;
      ModbusStatus : Word;
      A1_Scenario_Type : Int := 2;
      A2_Scenario_Type : Int := 1;
      B1_Scenario_Type : Int := 1;
      B2_Scenario_Type : Int := 1;
      A_Emergency : Bool;
      B_Emergency : Bool;
      A1_Fault : Bool;
      A2_Fault : Bool;
      B1_Fault : Bool;
      B2_Fault : Bool;
      A3_Fault : Bool;
      B3_Fault : Bool;
      A1_Silo_Low : Bool;
      A2_Silo_Low : Bool;
      B1_Silo_Low : Bool;
      B2_Silo_Low : Bool;
      A1_Conveyer : Bool;
      A2_Conveyer : Bool;
      B1_Conveyer : Bool;
      B2_Conveyer : Bool;
      A3_Conveyor : Bool;
      B3_Left_Conveyer : Bool;
      A1_Silo_High : Bool;
      A2_Silo_High : Bool;
      B1_Silo_High : Bool;
      B2_Silo_High : Bool;
      A1_Sample : Bool;
      A2_Sample : Bool;
      B1_Sample : Bool;
      B2_Sample : Bool;
      A1_Running_Duration : Time;
      A1_Pause_Duration : Time;
      A1_Feeder_Vibration_Intensity : Int;
      A1_Ruuning_Online : Time;
      A1_Pause_Online : Time;
      A1_Sample_Interval : Time;
      A1_Sample_Duration : Time;
      A1_Sample_Online : Time;
      A1_Enable : Bool;
      A1_Start : Bool;
      A1_Big_Silo : Bool;
      B1_Running_Duration : Time;
      B1_Pause_Duration : Time;
      B1_Feeder_Vibration_Intensity : Int;
      B1_Ruuning_Online : Time;
      B1_Pause_Online : Time;
      B1_Sample_Interval : Time;
      B1_Sample_Duration : Time;
      B1_Sample_Online : Time;
      B1_Enable : Bool;
      B1_Start : Bool;
      B1_Big_Silo : Bool;
      A2_Running_Duration : Time;
      A2_Pause_Duration : Time;
      A2_Feeder_Vibration_Intensity : Int;
      A2_Ruuning_Online : Time;
      A2_Pause_Online : Time;
      A2_Sample_Interval : Time;
      A2_Sample_Duration : Time;
      A2_Sample_Online : Time;
      A2_Enable : Bool;
      A2_Start : Bool;
      A2_Big_Silo : Bool;
      B2_Running_Duration : Time;
      B2_Pause_Duration : Time;
      B2_Feeder_Vibration_Intensity : Int;
      B2_Ruuning_Online : Time;
      B2_Pause_Online : Time;
      B2_Sample_Interval : Time;
      B2_Sample_Duration : Time;
      B2_Sample_Online : Time;
      B2_Enable : Bool;
      B2_Start : Bool;
      B2_Big_Silo : Bool;
      A1_Manual : Bool;
      A2_Manual : Bool;
      B1_Manual : Bool;
      B2_Manual : Bool;
      A1_Feeder : Bool;
      A2_Feeder : Bool;
      B1_Feeder : Bool;
      B2_Feeder : Bool;
      A1_Duration_Big_Silo_Stop_Time : Time;
      A2_Duration_Big_Silo_Stop_Time : Time;
      B1_Duration_Big_Silo_Stop_Time : Time;
      B2_Duration_Big_Silo_Stop_Time : Time;
      A1_Empty_Line_Time : Time;
      A2_Empty_Line_Time : Time;
      B1_Empty_Line_Time : Time;
      B2_Empty_Line_Time : Time;
      A1_Feeder_Delay_After_Start_Time : Time;
      A2_Feeder_Delay_After_Start_Time : Time;
      B1_Feeder_Delay_After_Start_Time : Time;
      B2_Feeder_Delay_After_Start_Time : Time;
      A1_Feeder_Delay_Before_Stop_Time : Time;
      A2_Feeder_Delay_Before_Stop_Time : Time;
      B1_Feeder_Delay_Before_Stop_Time : Time;
      B2_Feeder_Delay_Before_Stop_Time : Time;
      A1_Feeder_Delay_Time : Time;
      A1_Feeder_Delay_Time_1 : Time;
      A1_Feeder_Delay_Time_2 : Time;
      A1_Feeder_Delay_Time_3 : Time;
      B3_Conveyor : Bool;
   END_VAR
BEGIN
END_DATA_BLOCK

DATA_BLOCK "ConveyerA3_B3_DB"   // DB32
{ S7_Optimized_Access := 'TRUE' }
VERSION : 0.1
// stored: InstanceOfName ConveyerA3_B3
"ConveyerA3_B3"
BEGIN
END_DATA_BLOCK

DATA_BLOCK "Sample_A_DB"   // DB33
{ S7_Optimized_Access := 'TRUE' }
VERSION : 0.1
// stored: InstanceOfName Sample
"Sample"
BEGIN
END_DATA_BLOCK

DATA_BLOCK "Silo_Big_A-B_DB"   // DB34
{ S7_Optimized_Access := 'TRUE' }
VERSION : 0.1
// stored: InstanceOfName Silo_Big_A-B
"Silo_Big_A-B"
BEGIN
END_DATA_BLOCK

DATA_BLOCK "Web_Recieve"   // DB45
{ S7_Optimized_Access := 'FALSE' }